// TIA Portal project "Mes_Con" (V17) (continued)
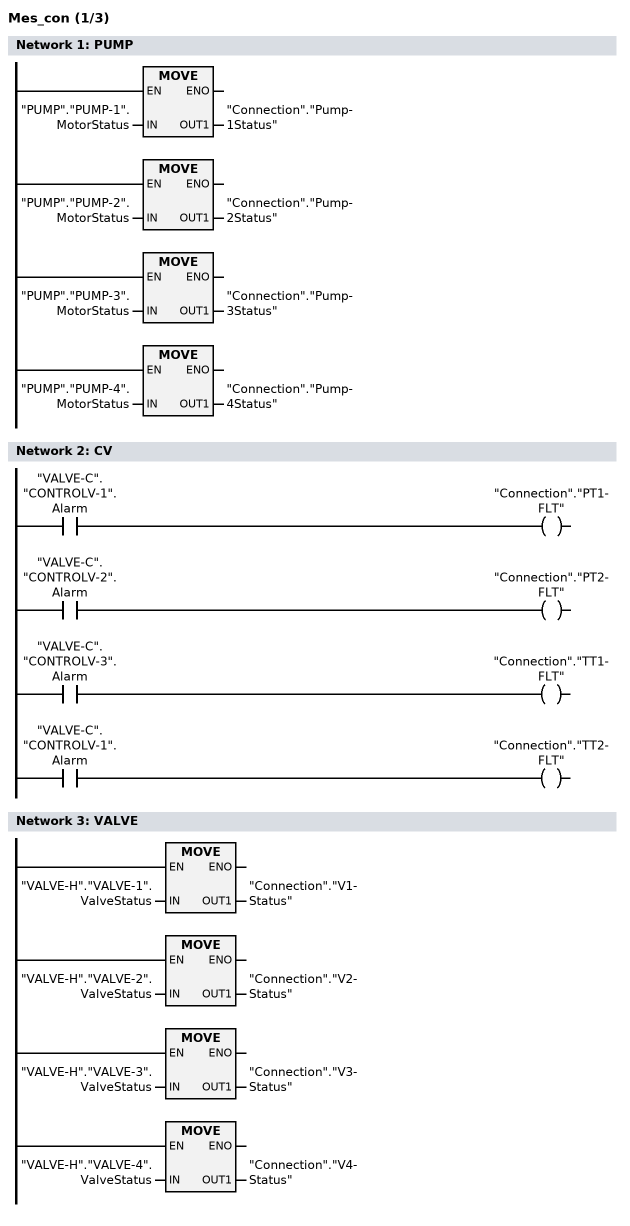
   RUNG wire#powerrail
      Move(in := "PUMP"."PUMP-1".MotorStatus, out1 => "Connection"."Pump-1Status")
   END_RUNG
   RUNG wire#powerrail
      Move(in := "PUMP"."PUMP-2".MotorStatus, out1 => "Connection"."Pump-2Status")
   END_RUNG
   RUNG wire#powerrail
      Move(in := "PUMP"."PUMP-3".MotorStatus, out1 => "Connection"."Pump-3Status")
   END_RUNG
   RUNG wire#powerrail
      Move(in := "PUMP"."PUMP-4".MotorStatus, out1 => "Connection"."Pump-4Status")
   END_RUNG
   // the same network as SCL:
   "Connection"."Pump-1Status" := "PUMP"."PUMP-1".MotorStatus;
   "Connection"."Pump-2Status" := "PUMP"."PUMP-2".MotorStatus;
   "Connection"."Pump-3Status" := "PUMP"."PUMP-3".MotorStatus;
   "Connection"."Pump-4Status" := "PUMP"."PUMP-4".MotorStatus;
END_REGION

REGION Network 2: CV
   RUNG wire#powerrail
      Contact( "VALVE-C"."CONTROLV-1".Alarm )
      Coil( "Connection"."PT1-FLT" )
   END_RUNG
   RUNG wire#powerrail
      Contact( "VALVE-C"."CONTROLV-2".Alarm )
      Coil( "Connection"."PT2-FLT" )
   END_RUNG
   RUNG wire#powerrail
      Contact( "VALVE-C"."CONTROLV-3".Alarm )
      Coil( "Connection"."TT1-FLT" )
   END_RUNG
   RUNG wire#powerrail
      Contact( "VALVE-C"."CONTROLV-1".Alarm )
      Coil( "Connection"."TT2-FLT" )
   END_RUNG
   // the same network as SCL:
   "Connection"."PT1-FLT" := "VALVE-C"."CONTROLV-1".Alarm;
   "Connection"."PT2-FLT" := "VALVE-C"."CONTROLV-2".Alarm;
   "Connection"."TT1-FLT" := "VALVE-C"."CONTROLV-3".Alarm;
   "Connection"."TT2-FLT" := "VALVE-C"."CONTROLV-1".Alarm;
END_REGION

REGION Network 3: VALVE
   RUNG wire#powerrail
      Move(in := "VALVE-H"."VALVE-1".ValveStatus, out1 => "Connection"."V1-Status")
   END_RUNG
   RUNG wire#powerrail
      Move(in := "VALVE-H"."VALVE-2".ValveStatus, out1 => "Connection"."V2-Status")
   END_RUNG
   RUNG wire#powerrail
      Move(in := "VALVE-H"."VALVE-3".ValveStatus, out1 => "Connection"."V3-Status")
   END_RUNG
   RUNG wire#powerrail
      Move(in := "VALVE-H"."VALVE-4".ValveStatus, out1 => "Connection"."V4-Status")
   END_RUNG
   // the same network as SCL:
   "Connection"."V1-Status" := "VALVE-H"."VALVE-1".ValveStatus;
   "Connection"."V2-Status" := "VALVE-H"."VALVE-2".ValveStatus;
   "Connection"."V3-Status" := "VALVE-H"."VALVE-3".ValveStatus;
   "Connection"."V4-Status" := "VALVE-H"."VALVE-4".ValveStatus;
END_REGION

REGION Network 4: TT
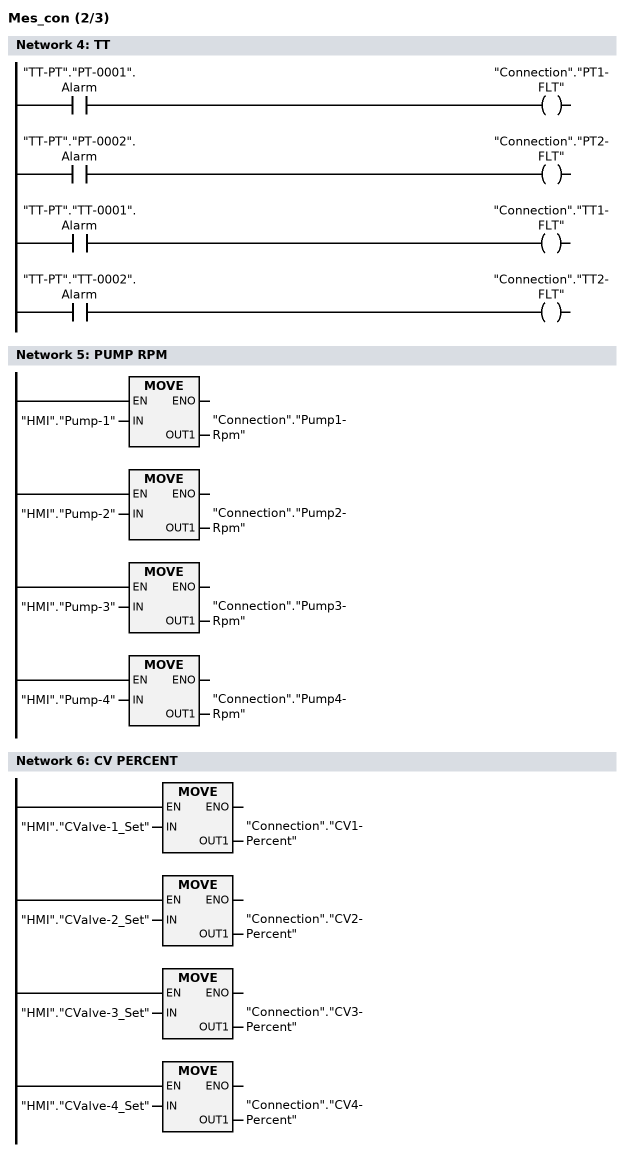
   RUNG wire#powerrail
      Contact( "TT-PT"."PT-0001".Alarm )
      Coil( "Connection"."PT1-FLT" )
   END_RUNG
   RUNG wire#powerrail
      Contact( "TT-PT"."PT-0002".Alarm )
      Coil( "Connection"."PT2-FLT" )
   END_RUNG
   RUNG wire#powerrail
      Contact( "TT-PT"."TT-0001".Alarm )
      Coil( "Connection"."TT1-FLT" )
   END_RUNG
   RUNG wire#powerrail
      Contact( "TT-PT"."TT-0002".Alarm )
      Coil( "Connection"."TT2-FLT" )
   END_RUNG
   // the same network as SCL:
   "Connection"."PT1-FLT" := "TT-PT"."PT-0001".Alarm;
   "Connection"."PT2-FLT" := "TT-PT"."PT-0002".Alarm;
   "Connection"."TT1-FLT" := "TT-PT"."TT-0001".Alarm;
   "Connection"."TT2-FLT" := "TT-PT"."TT-0002".Alarm;
END_REGION

REGION Network 5: PUMP RPM
   RUNG wire#powerrail
      Move(in := "HMI"."Pump-1", out1 => "Connection"."Pump1-Rpm")
   END_RUNG
   RUNG wire#powerrail
      Move(in := "HMI"."Pump-2", out1 => "Connection"."Pump2-Rpm")
   END_RUNG
   RUNG wire#powerrail
      Move(in := "HMI"."Pump-3", out1 => "Connection"."Pump3-Rpm")
   END_RUNG
   RUNG wire#powerrail
      Move(in := "HMI"."Pump-4", out1 => "Connection"."Pump4-Rpm")
   END_RUNG
   // the same network as SCL:
   "Connection"."Pump1-Rpm" := "HMI"."Pump-1";
   "Connection"."Pump2-Rpm" := "HMI"."Pump-2";
   "Connection"."Pump3-Rpm" := "HMI"."Pump-3";
   "Connection"."Pump4-Rpm" := "HMI"."Pump-4";
END_REGION

REGION Network 6: CV PERCENT
   RUNG wire#powerrail
      Move(in := "HMI"."CValve-1_Set", out1 => "Connection"."CV1-Percent")
   END_RUNG
   RUNG wire#powerrail
      Move(in := "HMI"."CValve-2_Set", out1 => "Connection"."CV2-Percent")
   END_RUNG
   RUNG wire#powerrail
      Move(in := "HMI"."CValve-3_Set", out1 => "Connection"."CV3-Percent")
   END_RUNG
   RUNG wire#powerrail
      Move(in := "HMI"."CValve-4_Set", out1 => "Connection"."CV4-Percent")
   END_RUNG
   // the same network as SCL:
   "Connection"."CV1-Percent" := "HMI"."CValve-1_Set";
   "Connection"."CV2-Percent" := "HMI"."CValve-2_Set";
   "Connection"."CV3-Percent" := "HMI"."CValve-3_Set";
   "Connection"."CV4-Percent" := "HMI"."CValve-4_Set";
END_REGION

REGION Network 7: ANOLOG VALUE
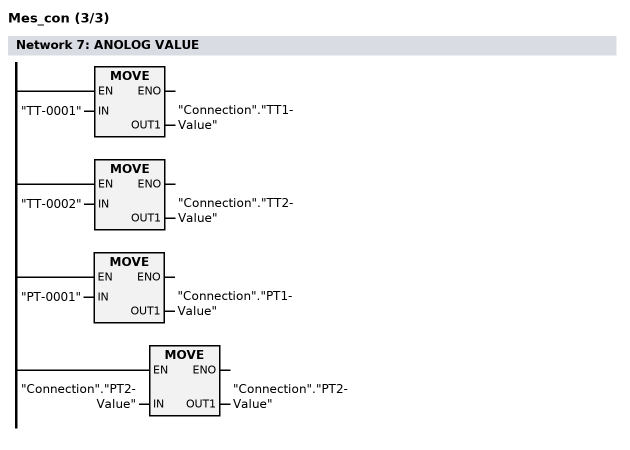
   RUNG wire#powerrail
      Move(in := "TT-0001", out1 => "Connection"."TT1-Value")
   END_RUNG
   RUNG wire#powerrail
      Move(in := "TT-0002", out1 => "Connection"."TT2-Value")
   END_RUNG
   RUNG wire#powerrail
      Move(in := "PT-0001", out1 => "Connection"."PT1-Value")
   END_RUNG
   RUNG wire#powerrail
      Move(in := "Connection"."PT2-Value", out1 => "Connection"."PT2-Value")
   END_RUNG
   // the same network as SCL:
   "Connection"."TT1-Value" := "TT-0001";
   "Connection"."TT2-Value" := "TT-0002";
   "Connection"."PT1-Value" := "PT-0001";
   "Connection"."PT2-Value" := "Connection"."PT2-Value";
END_REGION
END_FUNCTION

// folder: Eqp

FUNCTION "fncEl_VanasI" : Void   // FC6, LAD
{ S7_Optimized_Access := 'TRUE' }
VERSION : 0.1
   VAR_INPUT
      Vana_Opened : Bool;
      Vana_Closed : Bool;
      TımeOut : Int;
   END_VAR
   VAR_OUTPUT
      Alm : Bool;
      TWO_SIGNAL : Bool;
      NOT_SIGNAL : Bool;
   END_VAR
   VAR_IN_OUT
      ElVanası : "ElValve";
   END_VAR
   VAR_TEMP   // added for the SCL form of the ladder/FBD networks
      _w1 : Bool;
      _w2 : Bool;
   END_VAR
BEGIN

REGION Network 1: ATAMA
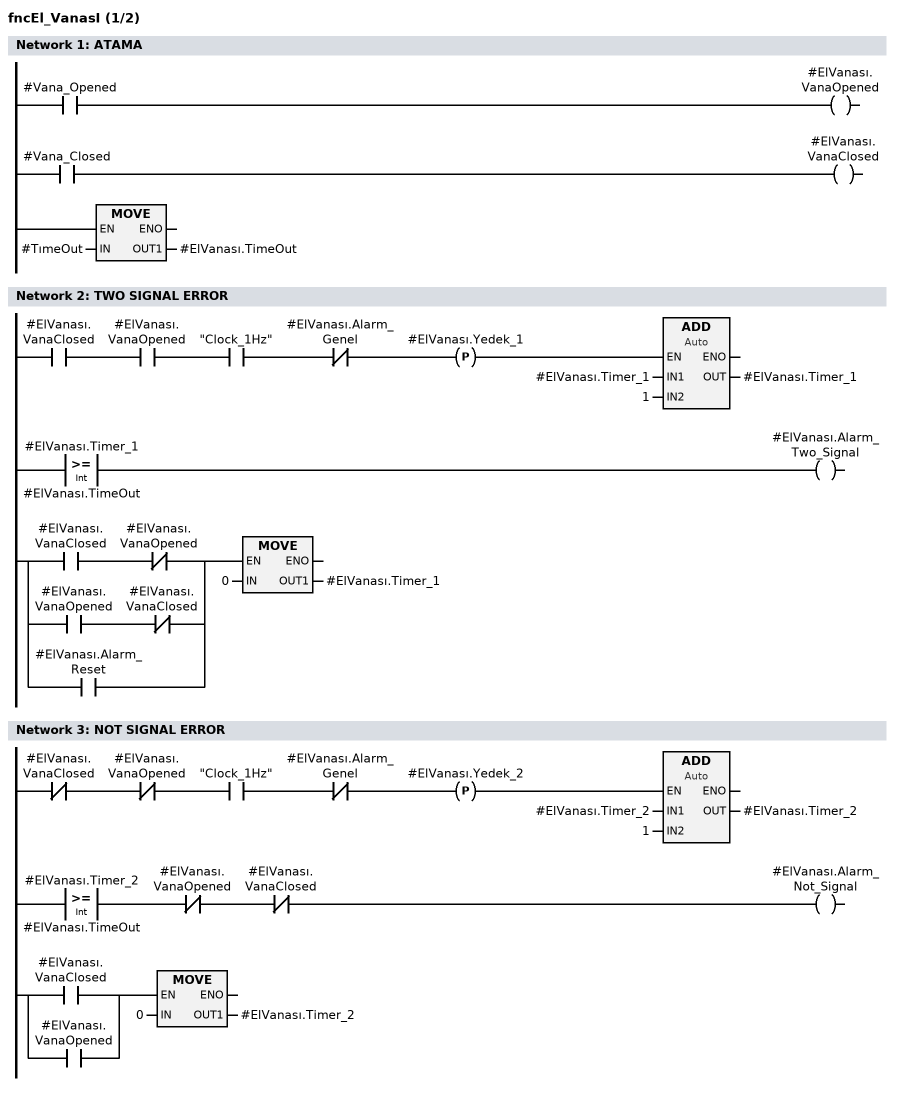
   RUNG wire#powerrail
      Contact( #Vana_Opened )
      Coil( #ElVanası.VanaOpened )
   END_RUNG
   RUNG wire#powerrail
      Contact( #Vana_Closed )
      Coil( #ElVanası.VanaClosed )
   END_RUNG
   RUNG wire#powerrail
      Move(in := #TımeOut, out1 => #ElVanası.TimeOut)
   END_RUNG
   // the same network as SCL:
   #ElVanası.VanaOpened := #Vana_Opened;
   #ElVanası.VanaClosed := #Vana_Closed;
   #ElVanası.TimeOut := #TımeOut;
END_REGION

REGION Network 2: TWO SIGNAL ERROR
   RUNG wire#powerrail
      Contact( #ElVanası.VanaClosed )
      Contact( #ElVanası.VanaOpened )
      Contact( "Clock_1Hz" )
      I_Contact( #ElVanası.Alarm_Genel )
      P_Trig( #ElVanası.Yedek_1 )
      Add(in1 := #ElVanası.Timer_1, in2 := 1, out => #ElVanası.Timer_1)
   END_RUNG
   RUNG wire#powerrail
      { S7_Templates := "SrcType := Int" } GE_Contact(in1 := #ElVanası.Timer_1, in2 := #ElVanası.TimeOut)
      Coil( #ElVanası.Alarm_Two_Signal )
   END_RUNG
   RUNG wire#powerrail
      Contact( #ElVanası.VanaClosed )
      I_Contact( #ElVanası.VanaOpened )
      wire#w1
      Move(in := 0, out1 => #ElVanası.Timer_1)
   END_RUNG
   RUNG wire#powerrail
      Contact( #ElVanası.VanaOpened )
      I_Contact( #ElVanası.VanaClosed )
   END_RUNG wire#w1
   RUNG wire#powerrail
      Contact( #ElVanası.Alarm_Reset )
   END_RUNG wire#w1
   // the same network as SCL:
   #_w1 := #ElVanası.VanaClosed AND #ElVanası.VanaOpened AND "Clock_1Hz" AND NOT #ElVanası.Alarm_Genel;
   #_w2 := #_w1 AND NOT #ElVanası.Yedek_1;   // rising edge
   #ElVanası.Yedek_1 := #_w1;
   IF #_w2 THEN #ElVanası.Timer_1 := #ElVanası.Timer_1 + 1; END_IF;
   #ElVanası.Alarm_Two_Signal := #ElVanası.Timer_1 >= #ElVanası.TimeOut;
   IF (#ElVanası.VanaClosed AND NOT #ElVanası.VanaOpened) OR (#ElVanası.VanaOpened AND NOT #ElVanası.VanaClosed) OR #ElVanası.Alarm_Reset THEN
       #ElVanası.Timer_1 := 0;
   END_IF;
END_REGION

REGION Network 3: NOT SIGNAL ERROR
   RUNG wire#powerrail
      I_Contact( #ElVanası.VanaClosed )
      I_Contact( #ElVanası.VanaOpened )
      Contact( "Clock_1Hz" )
      I_Contact( #ElVanası.Alarm_Genel )
      P_Trig( #ElVanası.Yedek_2 )
      Add(in1 := #ElVanası.Timer_2, in2 := 1, out => #ElVanası.Timer_2)
   END_RUNG
   RUNG wire#powerrail
      { S7_Templates := "SrcType := Int" } GE_Contact(in1 := #ElVanası.Timer_2, in2 := #ElVanası.TimeOut)
      I_Contact( #ElVanası.VanaOpened )
      I_Contact( #ElVanası.VanaClosed )
      Coil( #ElVanası.Alarm_Not_Signal )
   END_RUNG
   RUNG wire#powerrail
      Contact( #ElVanası.VanaClosed )
      wire#w1
      Move(in := 0, out1 => #ElVanası.Timer_2)
   END_RUNG
   RUNG wire#powerrail
      Contact( #ElVanası.VanaOpened )
   END_RUNG wire#w1
   // the same network as SCL:
   #_w1 := NOT #ElVanası.VanaClosed AND NOT #ElVanası.VanaOpened AND "Clock_1Hz" AND NOT #ElVanası.Alarm_Genel;
   #_w2 := #_w1 AND NOT #ElVanası.Yedek_2;   // rising edge
   #ElVanası.Yedek_2 := #_w1;
   IF #_w2 THEN #ElVanası.Timer_2 := #ElVanası.Timer_2 + 1; END_IF;
   #ElVanası.Alarm_Not_Signal := (#ElVanası.Timer_2 >= #ElVanası.TimeOut) AND NOT #ElVanası.VanaOpened AND NOT #ElVanası.VanaClosed;
   IF #ElVanası.VanaClosed OR #ElVanası.VanaOpened THEN #ElVanası.Timer_2 := 0; END_IF;
END_REGION

REGION Network 4: GENEL ALARM
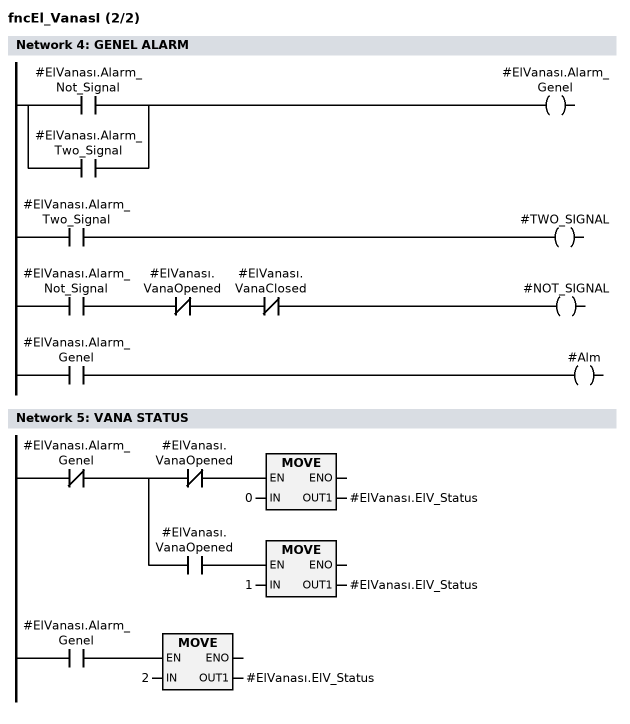
   RUNG wire#powerrail
      Contact( #ElVanası.Alarm_Not_Signal )
      wire#w1
      Coil( #ElVanası.Alarm_Genel )
   END_RUNG
   RUNG wire#powerrail
      Contact( #ElVanası.Alarm_Two_Signal )
   END_RUNG wire#w1
   RUNG wire#powerrail
      Contact( #ElVanası.Alarm_Two_Signal )
      Coil( #TWO_SIGNAL )
   END_RUNG
   RUNG wire#powerrail
      Contact( #ElVanası.Alarm_Not_Signal )
      I_Contact( #ElVanası.VanaOpened )
      I_Contact( #ElVanası.VanaClosed )
      Coil( #NOT_SIGNAL )
   END_RUNG
   RUNG wire#powerrail
      Contact( #ElVanası.Alarm_Genel )
      Coil( #Alm )
   END_RUNG
   // the same network as SCL:
   #ElVanası.Alarm_Genel := #ElVanası.Alarm_Not_Signal OR #ElVanası.Alarm_Two_Signal;
   #TWO_SIGNAL := #ElVanası.Alarm_Two_Signal;
   #NOT_SIGNAL := #ElVanası.Alarm_Not_Signal AND NOT #ElVanası.VanaOpened AND NOT #ElVanası.VanaClosed;
   #Alm := #ElVanası.Alarm_Genel;
END_REGION

REGION Network 5: VANA STATUS
   RUNG wire#powerrail
      I_Contact( #ElVanası.Alarm_Genel )
      wire#w1
      I_Contact( #ElVanası.VanaOpened )
      Move(in := 0, out1 => #ElVanası.ElV_Status)
   END_RUNG
   RUNG wire#w1
      Contact( #ElVanası.VanaOpened )
      Move(in := 1, out1 => #ElVanası.ElV_Status)
   END_RUNG
   RUNG wire#powerrail
      Contact( #ElVanası.Alarm_Genel )
      Move(in := 2, out1 => #ElVanası.ElV_Status)
   END_RUNG
   // the same network as SCL:
   #_w1 := NOT #ElVanası.Alarm_Genel;
   IF #_w1 AND NOT #ElVanası.VanaOpened THEN #ElVanası.ElV_Status := 0; END_IF;
   IF #_w1 AND #ElVanası.VanaOpened THEN #ElVanası.ElV_Status := 1; END_IF;
   IF #ElVanası.Alarm_Genel THEN #ElVanası.ElV_Status := 2; END_IF;
END_REGION
END_FUNCTION

FUNCTION "fncFlow" : Void   // FC13, LAD
{ S7_Optimized_Access := 'TRUE' }
VERSION : 0.1
   VAR_INPUT
      Pulse : Bool;
      FwValue : Real;
      Pulse_Kg : Real;
      Reset : Bool;
      TankBoşaltıldı : Bool;
      Tank_Valur_reset : Bool;
      Su_Alım_Run : Bool;
      inflight : DInt;
   END_VAR
   VAR_IN_OUT
      FM : "FM";
   END_VAR
   VAR_TEMP   // added for the SCL form of the ladder/FBD networks
      _w1 : Bool;
   END_VAR
BEGIN

REGION Network 1: Atama
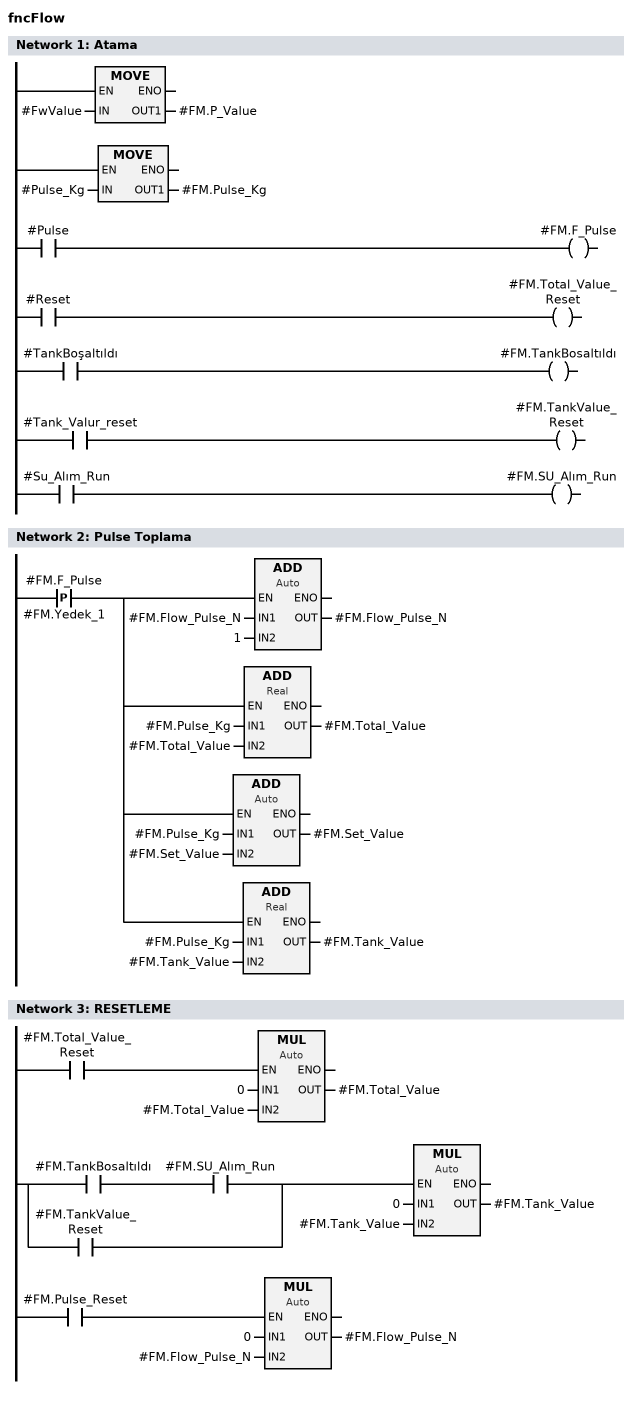
   RUNG wire#powerrail
      Move(in := #FwValue, out1 => #FM.P_Value)
   END_RUNG
   RUNG wire#powerrail
      Move(in := #Pulse_Kg, out1 => #FM.Pulse_Kg)
   END_RUNG
   RUNG wire#powerrail
      Contact( #Pulse )
      Coil( #FM.F_Pulse )
   END_RUNG
   RUNG wire#powerrail
      Contact( #Reset )
      Coil( #FM.Total_Value_Reset )
   END_RUNG
   RUNG wire#powerrail
      Contact( #TankBoşaltıldı )
      Coil( #FM.TankBosaltıldı )
   END_RUNG
   RUNG wire#powerrail
      Contact( #Tank_Valur_reset )
      Coil( #FM.TankValue_Reset )
   END_RUNG
   RUNG wire#powerrail
      Contact( #Su_Alım_Run )
      Coil( #FM.SU_Alım_Run )
   END_RUNG
   // the same network as SCL:
   #FM.P_Value := #FwValue;
   #FM.Pulse_Kg := #Pulse_Kg;
   #FM.F_Pulse := #Pulse;
   #FM.Total_Value_Reset := #Reset;
   #FM.TankBosaltıldı := #TankBoşaltıldı;
   #FM.TankValue_Reset := #Tank_Valur_reset;
   #FM.SU_Alım_Run := #Su_Alım_Run;
END_REGION

REGION Network 2: Pulse Toplama
   RUNG wire#powerrail
      P_Contact(operand := #FM.F_Pulse, bit := #FM.Yedek_1)
      wire#w1
      Add(in1 := #FM.Flow_Pulse_N, in2 := 1, out => #FM.Flow_Pulse_N)
   END_RUNG
   RUNG wire#w1
      { S7_Templates := "SrcType := Real" } Add(in1 := #FM.Pulse_Kg, in2 := #FM.Total_Value, out => #FM.Total_Value)
   END_RUNG
   RUNG wire#w1
      Add(in1 := #FM.Pulse_Kg, in2 := #FM.Set_Value, out => #FM.Set_Value)
   END_RUNG
   RUNG wire#w1
      { S7_Templates := "SrcType := Real" } Add(in1 := #FM.Pulse_Kg, in2 := #FM.Tank_Value, out => #FM.Tank_Value)
   END_RUNG
   // the same network as SCL:
   #_w1 := #FM.F_Pulse AND NOT #FM.Yedek_1;   // rising edge of #FM.F_Pulse
   #FM.Yedek_1 := #FM.F_Pulse;
   IF #_w1 THEN
       #FM.Flow_Pulse_N := #FM.Flow_Pulse_N + 1;
       #FM.Total_Value := #FM.Pulse_Kg + #FM.Total_Value;
       #FM.Set_Value := #FM.Pulse_Kg + #FM.Set_Value;
       #FM.Tank_Value := #FM.Pulse_Kg + #FM.Tank_Value;
   END_IF;
END_REGION

REGION Network 3: RESETLEME
   RUNG wire#powerrail
      Contact( #FM.Total_Value_Reset )
      Mul(in1 := 0, in2 := #FM.Total_Value, out => #FM.Total_Value)
   END_RUNG
   RUNG wire#powerrail
      Contact( #FM.TankBosaltıldı )
      Contact( #FM.SU_Alım_Run )
      wire#w1
      Mul(in1 := 0, in2 := #FM.Tank_Value, out => #FM.Tank_Value)
   END_RUNG
   RUNG wire#powerrail
      Contact( #FM.TankValue_Reset )
   END_RUNG wire#w1
   RUNG wire#powerrail
      Contact( #FM.Pulse_Reset )
      Mul(in1 := 0, in2 := #FM.Flow_Pulse_N, out => #FM.Flow_Pulse_N)
   END_RUNG
   // the same network as SCL:
   IF #FM.Total_Value_Reset THEN #FM.Total_Value := 0 * #FM.Total_Value; END_IF;
   IF (#FM.TankBosaltıldı AND #FM.SU_Alım_Run) OR #FM.TankValue_Reset THEN
       #FM.Tank_Value := 0 * #FM.Tank_Value;
   END_IF;
   IF #FM.Pulse_Reset THEN #FM.Flow_Pulse_N := 0 * #FM.Flow_Pulse_N; END_IF;
END_REGION
END_FUNCTION

// folder: Eqp/Anolog

FUNCTION "fncAI" : Void   // FC5, LAD
{ S7_Optimized_Access := 'TRUE' }
VERSION : 0.1
   VAR_INPUT
      Analog_Input : Int;
   END_VAR
   VAR_OUTPUT
      Alarm : Bool;
   END_VAR
   VAR_IN_OUT
      "A" : "AnalogInput";
   END_VAR
   VAR_TEMP   // added for the SCL form of the ladder/FBD networks
      _w1 : Bool;
      _w2 : Bool;
   END_VAR
BEGIN

REGION Network 1: ATAMA
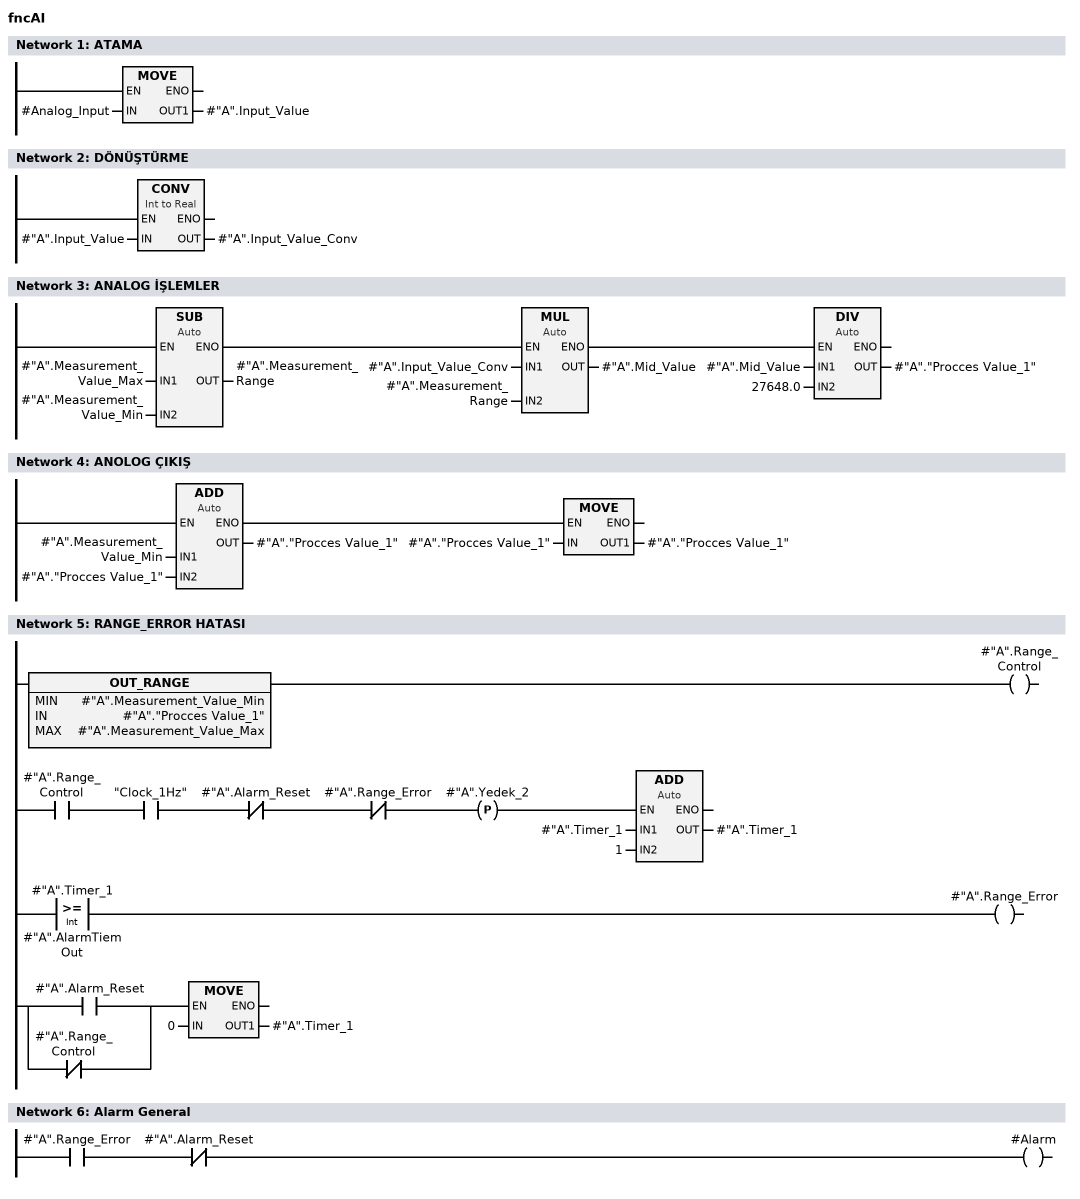
   RUNG wire#powerrail
      Move(in := #Analog_Input, out1 => #"A".Input_Value)
   END_RUNG
   // the same network as SCL:
   #"A".Input_Value := #Analog_Input;
END_REGION

REGION Network 2: DÖNÜŞTÜRME
   RUNG wire#powerrail
      { S7_Templates := "[SrcType := Int, DestType := Real]" } Convert(in := #"A".Input_Value, out => #"A".Input_Value_Conv)
   END_RUNG
   // the same network as SCL:
   #"A".Input_Value_Conv := INT_TO_REAL(#"A".Input_Value);
END_REGION

REGION Network 3: ANALOG İŞLEMLER
   RUNG wire#powerrail
      Sub(in1 := #"A".Measurement_Value_Max, in2 := #"A".Measurement_Value_Min, out => #"A".Measurement_Range)
      Mul(in1 := #"A".Input_Value_Conv, in2 := #"A".Measurement_Range, out => #"A".Mid_Value)
      Div(in1 := #"A".Mid_Value, in2 := 27648.0, out => #"A"."Procces Value_1")
   END_RUNG
   // the same network as SCL:
   #"A".Measurement_Range := #"A".Measurement_Value_Max - #"A".Measurement_Value_Min;
   #"A".Mid_Value := #"A".Input_Value_Conv * #"A".Measurement_Range;
   #"A"."Procces Value_1" := #"A".Mid_Value / 27648.0;
END_REGION

REGION Network 4: ANOLOG ÇIKIŞ
   RUNG wire#powerrail
      Add(in1 := #"A".Measurement_Value_Min, in2 := #"A"."Procces Value_1", out => #"A"."Procces Value_1")
      Move(in := #"A"."Procces Value_1", out1 => #"A"."Procces Value_1")
   END_RUNG
   // the same network as SCL:
   #"A"."Procces Value_1" := #"A".Measurement_Value_Min + #"A"."Procces Value_1";
   #"A"."Procces Value_1" := #"A"."Procces Value_1";
END_REGION

REGION Network 5: RANGE_ERROR HATASI
   #"A".Range_Control := (#"A"."Procces Value_1" < #"A".Measurement_Value_Min) OR (#"A"."Procces Value_1" > #"A".Measurement_Value_Max);
   #_w1 := #"A".Range_Control AND "Clock_1Hz" AND NOT #"A".Alarm_Reset AND NOT #"A".Range_Error;
   #_w2 := #_w1 AND NOT #"A".Yedek_2;   // rising edge
   #"A".Yedek_2 := #_w1;
   IF #_w2 THEN #"A".Timer_1 := #"A".Timer_1 + 1; END_IF;
   #"A".Range_Error := #"A".Timer_1 >= #"A".AlarmTiemOut;
   IF #"A".Alarm_Reset OR NOT #"A".Range_Control THEN #"A".Timer_1 := 0; END_IF;
END_REGION

REGION Network 6: Alarm General
   RUNG wire#powerrail
      Contact( #"A".Range_Error )
      I_Contact( #"A".Alarm_Reset )
      Coil( #Alarm )
   END_RUNG
   // the same network as SCL:
   #Alarm := #"A".Range_Error AND NOT #"A".Alarm_Reset;
END_REGION
END_FUNCTION

FUNCTION "fncAO" : Void   // FC7, LAD
{ S7_Optimized_Access := 'TRUE' }
VERSION : 0.1
   VAR_INPUT
      "Procces Value" : Real;
   END_VAR
   VAR_OUTPUT
      Proces_Value_Input : Int;
      Alarm : Bool;
   END_VAR
   VAR_IN_OUT
      AO : "AnalogOutput";
      Popup_1 : Bool;
   END_VAR
   VAR_TEMP   // added for the SCL form of the ladder/FBD networks
      _w1 : Bool;
      _w2 : Bool;
   END_VAR
BEGIN

REGION Network 1: ATAMA
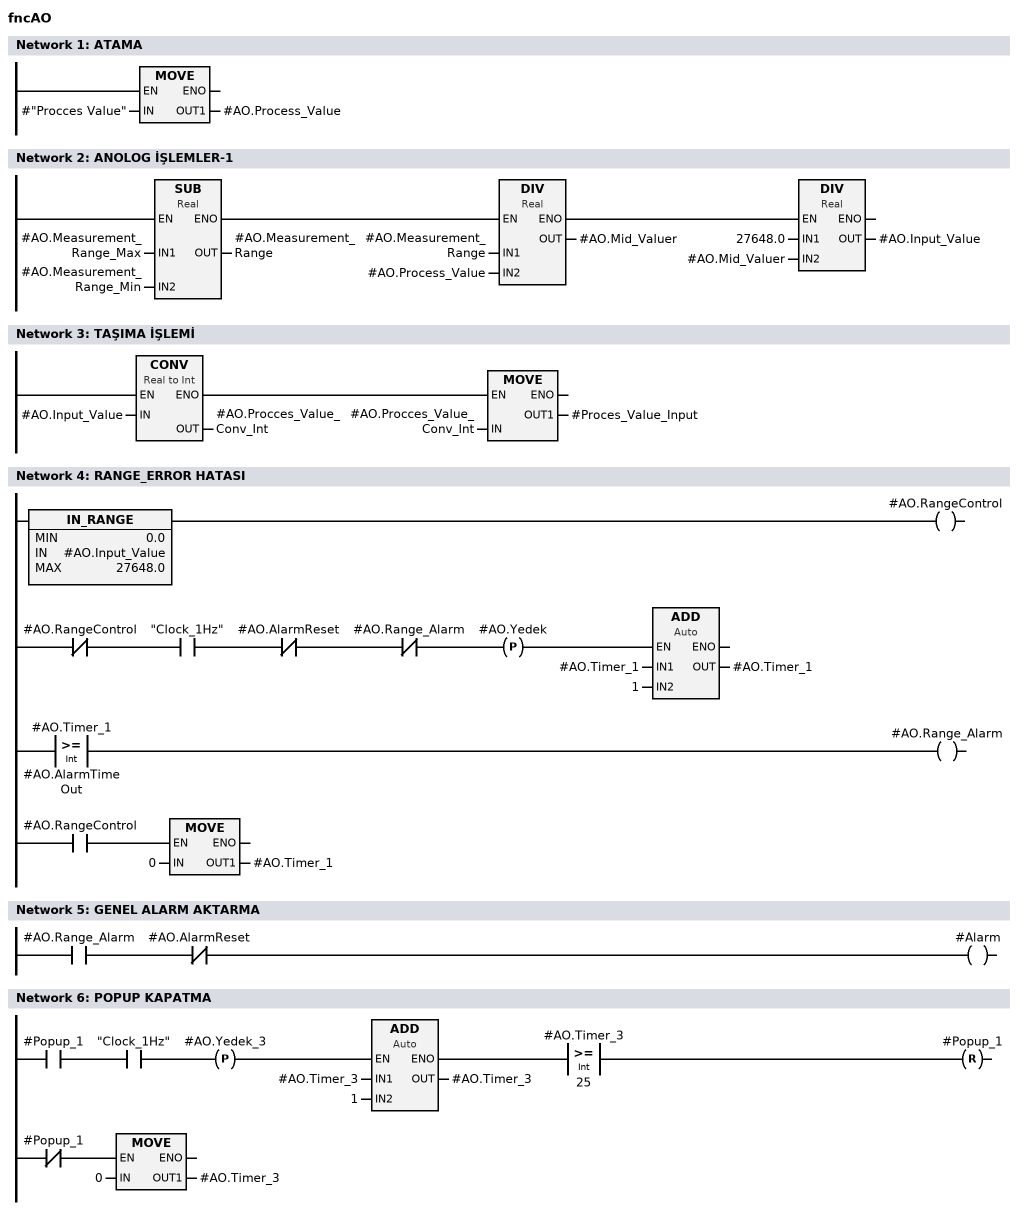
   RUNG wire#powerrail
      Move(in := #"Procces Value", out1 => #AO.Process_Value)
   END_RUNG
   // the same network as SCL:
   #AO.Process_Value := #"Procces Value";
END_REGION

REGION Network 2: ANOLOG İŞLEMLER-1
   RUNG wire#powerrail
      { S7_Templates := "SrcType := Real" } Sub(in1 := #AO.Measurement_Range_Max, in2 := #AO.Measurement_Range_Min, out => #AO.Measurement_Range)
      { S7_Templates := "SrcType := Real" } Div(in1 := #AO.Measurement_Range, in2 := #AO.Process_Value, out => #AO.Mid_Valuer)
      { S7_Templates := "SrcType := Real" } Div(in1 := 27648.0, in2 := #AO.Mid_Valuer, out => #AO.Input_Value)
   END_RUNG
   // the same network as SCL:
   #AO.Measurement_Range := #AO.Measurement_Range_Max - #AO.Measurement_Range_Min;
   #AO.Mid_Valuer := #AO.Measurement_Range / #AO.Process_Value;
   #AO.Input_Value := 27648.0 / #AO.Mid_Valuer;
END_REGION

REGION Network 3: TAŞIMA İŞLEMİ
   RUNG wire#powerrail
      { S7_Templates := "[SrcType := Real, DestType := Int]" } Convert(in := #AO.Input_Value, out => #AO.Procces_Value_Conv_Int)
      Move(in := #AO.Procces_Value_Conv_Int, out1 => #Proces_Value_Input)
   END_RUNG
   // the same network as SCL:
   #AO.Procces_Value_Conv_Int := REAL_TO_INT(#AO.Input_Value);
   #Proces_Value_Input := #AO.Procces_Value_Conv_Int;
END_REGION

REGION Network 4: RANGE_ERROR HATASI
   RUNG wire#powerrail
      { S7_Templates := "SrcType := Real" } InRange(min := 0.0, in := #AO.Input_Value, max := 27648.0)
      Coil( #AO.RangeControl )
   END_RUNG
   RUNG wire#powerrail
      I_Contact( #AO.RangeControl )
      Contact( "Clock_1Hz" )
      I_Contact( #AO.AlarmReset )
      I_Contact( #AO.Range_Alarm )
      P_Trig( #AO.Yedek )
      Add(in1 := #AO.Timer_1, in2 := 1, out => #AO.Timer_1)
   END_RUNG
   RUNG wire#powerrail
      { S7_Templates := "SrcType := Int" } GE_Contact(in1 := #AO.Timer_1, in2 := #AO.AlarmTimeOut)
      Coil( #AO.Range_Alarm )
   END_RUNG
   RUNG wire#powerrail
      Contact( #AO.RangeControl )
      Move(in := 0, out1 => #AO.Timer_1)
   END_RUNG
   // the same network as SCL:
   #AO.RangeControl := (0.0 <= #AO.Input_Value) AND (#AO.Input_Value <= 27648.0);
   #_w1 := NOT #AO.RangeControl AND "Clock_1Hz" AND NOT #AO.AlarmReset AND NOT #AO.Range_Alarm;
   #_w2 := #_w1 AND NOT #AO.Yedek;   // rising edge
   #AO.Yedek := #_w1;
   IF #_w2 THEN #AO.Timer_1 := #AO.Timer_1 + 1; END_IF;
   #AO.Range_Alarm := #AO.Timer_1 >= #AO.AlarmTimeOut;
   IF #AO.RangeControl THEN #AO.Timer_1 := 0; END_IF;
END_REGION

REGION Network 5: GENEL ALARM AKTARMA
   RUNG wire#powerrail
      Contact( #AO.Range_Alarm )
      I_Contact( #AO.AlarmReset )
      Coil( #Alarm )
   END_RUNG
   // the same network as SCL:
   #Alarm := #AO.Range_Alarm AND NOT #AO.AlarmReset;
END_REGION

REGION Network 6: POPUP KAPATMA
   RUNG wire#powerrail
      Contact( #Popup_1 )
      Contact( "Clock_1Hz" )
      P_Trig( #AO.Yedek_3 )
      Add(in1 := #AO.Timer_3, in2 := 1, out => #AO.Timer_3)
      { S7_Templates := "SrcType := Int" } GE_Contact(in1 := #AO.Timer_3, in2 := 25)
      R_Coil( #Popup_1 )
   END_RUNG
   RUNG wire#powerrail
      I_Contact( #Popup_1 )
      Move(in := 0, out1 => #AO.Timer_3)
   END_RUNG
   // the same network as SCL:
   #_w1 := #Popup_1 AND "Clock_1Hz";
   #_w2 := #_w1 AND NOT #AO.Yedek_3;   // rising edge
   #AO.Yedek_3 := #_w1;
   IF #_w2 THEN #AO.Timer_3 := #AO.Timer_3 + 1; END_IF;
   IF #_w2 AND (#AO.Timer_3 >= 25) THEN #Popup_1 := FALSE; END_IF;
   IF NOT #Popup_1 THEN #AO.Timer_3 := 0; END_IF;
END_REGION
END_FUNCTION

// folder: Eqp/Motor

FUNCTION "fncMotor" : Void   // FC1, LAD
{ S7_Optimized_Access := 'FALSE' }
VERSION : 0.1
   VAR_INPUT
      Mode : Bool;   // 0 = RunTime , 1 = Simulation
      MotorRunning : Bool;
      MotorThermic : Bool;
      Interlock : Bool;
      YU_Time : Int;
      MotorTimeOut : Int;
      "Local/Remote" : Bool;
   END_VAR
   VAR_OUTPUT
      "Motor Run" : Bool;
      ThermicAlarm : Bool;
      "M.TimeOut" : Bool;
      ShortCircuit : Bool;
      PhaseAlarm : Bool;
   END_VAR
   VAR_IN_OUT
      "M" : "Motor";
      Motor_Popup : Bool;
   END_VAR
   VAR_TEMP
      ALM : Struct
         ALM0 : Bool;
         ALM1 : Bool;
         ALM2 : Bool;
         ALM3 : Bool;
         ALM4 : Bool;
         ALM5 : Bool;
         ALM6 : Bool;
         ALM7 : Bool;
      END_STRUCT;
      temp : Bool;
      SimulationRUN : Bool;
   END_VAR
   VAR_TEMP   // added for the SCL form of the ladder/FBD networks
      _w1 : Bool;
      _w2 : Bool;
      _w3 : Bool;
      _w4 : Bool;
      _w5 : Bool;
      _w6 : Bool;
      _w7 : Bool;
   END_VAR
BEGIN

REGION Network 1: Input Atamaları
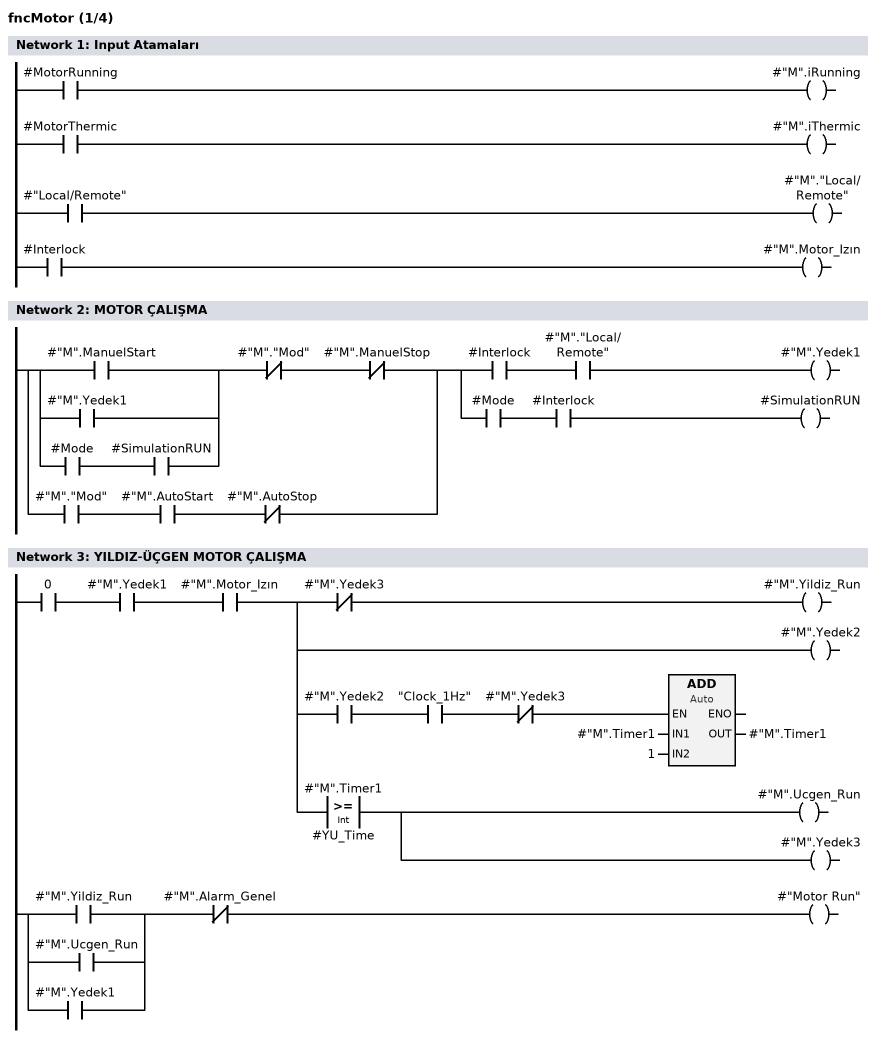
   RUNG wire#powerrail
      Contact( #MotorRunning )
      Coil( #"M".iRunning )
   END_RUNG
   RUNG wire#powerrail
      Contact( #MotorThermic )
      Coil( #"M".iThermic )
   END_RUNG
   RUNG wire#powerrail
      Contact( #"Local/Remote" )
      Coil( #"M"."Local/Remote" )
   END_RUNG
   RUNG wire#powerrail
      Contact( #Interlock )
      Coil( #"M".Motor_Izın )
   END_RUNG
   // the same network as SCL:
   #"M".iRunning := #MotorRunning;
   #"M".iThermic := #MotorThermic;
   #"M"."Local/Remote" := #"Local/Remote";
   #"M".Motor_Izın := #Interlock;
END_REGION

REGION Network 2: MOTOR ÇALIŞMA
   RUNG wire#powerrail
      Contact( #"M".ManuelStart )
      wire#w1
      I_Contact( #"M"."Mod" )
      I_Contact( #"M".ManuelStop )
      wire#w2
      Contact( #Interlock )
      Contact( #"M"."Local/Remote" )
      Coil( #"M".Yedek1 )
   END_RUNG
   RUNG wire#powerrail
      Contact( #"M".Yedek1 )
   END_RUNG wire#w1
   RUNG wire#powerrail
      Contact( #Mode )
      Contact( #SimulationRUN )
   END_RUNG wire#w1
   RUNG wire#powerrail
      Contact( #"M"."Mod" )
      Contact( #"M".AutoStart )
      I_Contact( #"M".AutoStop )
   END_RUNG wire#w2
   RUNG wire#w2
      Contact( #Mode )
      Contact( #Interlock )
      Coil( #SimulationRUN )
   END_RUNG
   // the same network as SCL:
   #_w1 := ((#"M".ManuelStart OR #"M".Yedek1 OR (#Mode AND #SimulationRUN)) AND NOT #"M"."Mod" AND NOT #"M".ManuelStop) OR (#"M"."Mod" AND #"M".AutoStart AND NOT #"M".AutoStop);
   #"M".Yedek1 := #_w1 AND #Interlock AND #"M"."Local/Remote";
   #SimulationRUN := #_w1 AND #Mode AND #Interlock;
END_REGION

REGION Network 3: YILDIZ-ÜÇGEN MOTOR ÇALIŞMA
   RUNG wire#powerrail
      Contact( 0 )
      Contact( #"M".Yedek1 )
      Contact( #"M".Motor_Izın )
      wire#w1
      I_Contact( #"M".Yedek3 )
      Coil( #"M".Yildiz_Run )
   END_RUNG
   RUNG wire#w1
      Coil( #"M".Yedek2 )
   END_RUNG
   RUNG wire#w1
      Contact( #"M".Yedek2 )
      Contact( "Clock_1Hz" )
      I_Contact( #"M".Yedek3 )
      Add(in1 := #"M".Timer1, in2 := 1, out => #"M".Timer1)
   END_RUNG
   RUNG wire#w1
      { S7_Templates := "SrcType := Int" } GE_Contact(in1 := #"M".Timer1, in2 := #YU_Time)
      wire#w2
      Coil( #"M".Ucgen_Run )
   END_RUNG
   RUNG wire#w2
      Coil( #"M".Yedek3 )
   END_RUNG
   RUNG wire#powerrail
      Contact( #"M".Yildiz_Run )
      wire#w3
      I_Contact( #"M".Alarm_Genel )
      Coil( #"Motor Run" )
   END_RUNG
   RUNG wire#powerrail
      Contact( #"M".Ucgen_Run )
   END_RUNG wire#w3
   RUNG wire#powerrail
      Contact( #"M".Yedek1 )
   END_RUNG wire#w3
   // the same network as SCL:
   #_w1 := 0 AND #"M".Yedek1 AND #"M".Motor_Izın;
   #"M".Yildiz_Run := #_w1 AND NOT #"M".Yedek3;
   #"M".Yedek2 := #_w1;
   IF #_w1 AND #"M".Yedek2 AND "Clock_1Hz" AND NOT #"M".Yedek3 THEN #"M".Timer1 := #"M".Timer1 + 1; END_IF;
   #"M".Ucgen_Run := #_w1 AND (#"M".Timer1 >= #YU_Time);
   #"M".Yedek3 := #"M".Ucgen_Run;
   #"Motor Run" := (#"M".Yildiz_Run OR #"M".Ucgen_Run OR #"M".Yedek1) AND NOT #"M".Alarm_Genel;
END_REGION

REGION Network 4: Motor Timeout Alarm
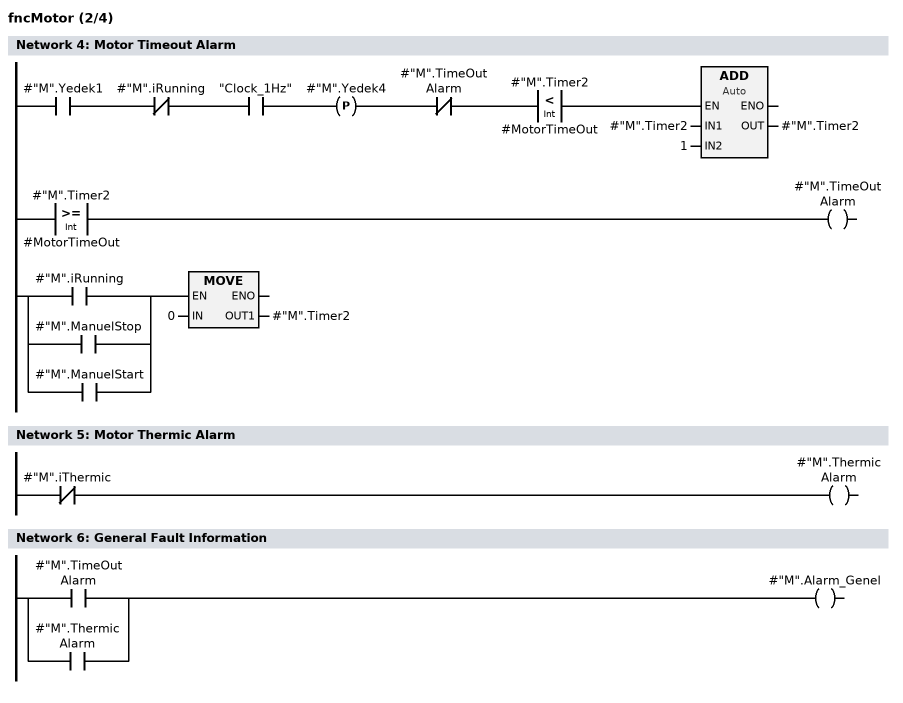
   RUNG wire#powerrail
      Contact( #"M".Yedek1 )
      I_Contact( #"M".iRunning )
      Contact( "Clock_1Hz" )
      P_Trig( #"M".Yedek4 )
      I_Contact( #"M".TimeOutAlarm )
      { S7_Templates := "SrcType := Int" } LT_Contact(in1 := #"M".Timer2, in2 := #MotorTimeOut)
      Add(in1 := #"M".Timer2, in2 := 1, out => #"M".Timer2)
   END_RUNG
   RUNG wire#powerrail
      { S7_Templates := "SrcType := Int" } GE_Contact(in1 := #"M".Timer2, in2 := #MotorTimeOut)
      Coil( #"M".TimeOutAlarm )
   END_RUNG
   RUNG wire#powerrail
      Contact( #"M".iRunning )
      wire#w1
      Move(in := 0, out1 => #"M".Timer2)
   END_RUNG
   RUNG wire#powerrail
      Contact( #"M".ManuelStop )
   END_RUNG wire#w1
   RUNG wire#powerrail
      Contact( #"M".ManuelStart )
   END_RUNG wire#w1
   // the same network as SCL:
   #_w1 := #"M".Yedek1 AND NOT #"M".iRunning AND "Clock_1Hz";
   #_w2 := #_w1 AND NOT #"M".Yedek4;   // rising edge
   #"M".Yedek4 := #_w1;
   IF #_w2 AND NOT #"M".TimeOutAlarm AND (#"M".Timer2 < #MotorTimeOut) THEN
       #"M".Timer2 := #"M".Timer2 + 1;
   END_IF;
   #"M".TimeOutAlarm := #"M".Timer2 >= #MotorTimeOut;
   IF #"M".iRunning OR #"M".ManuelStop OR #"M".ManuelStart THEN #"M".Timer2 := 0; END_IF;
END_REGION

REGION Network 5: Motor Thermic Alarm
   RUNG wire#powerrail
      I_Contact( #"M".iThermic )
      Coil( #"M".ThermicAlarm )
   END_RUNG
   // the same network as SCL:
   #"M".ThermicAlarm := NOT #"M".iThermic;
END_REGION

REGION Network 6: General Fault Information
   RUNG wire#powerrail
      Contact( #"M".TimeOutAlarm )
      wire#w1
      Coil( #"M".Alarm_Genel )
   END_RUNG
   RUNG wire#powerrail
      Contact( #"M".ThermicAlarm )
   END_RUNG wire#w1
   // the same network as SCL:
   #"M".Alarm_Genel := #"M".TimeOutAlarm OR #"M".ThermicAlarm;
END_REGION

REGION Network 7: Motor Status
   // 0 = Orjinal Rengi
   // 1 = Yeşil
   // 2 = Sarı
   // 3 = Kırmızı